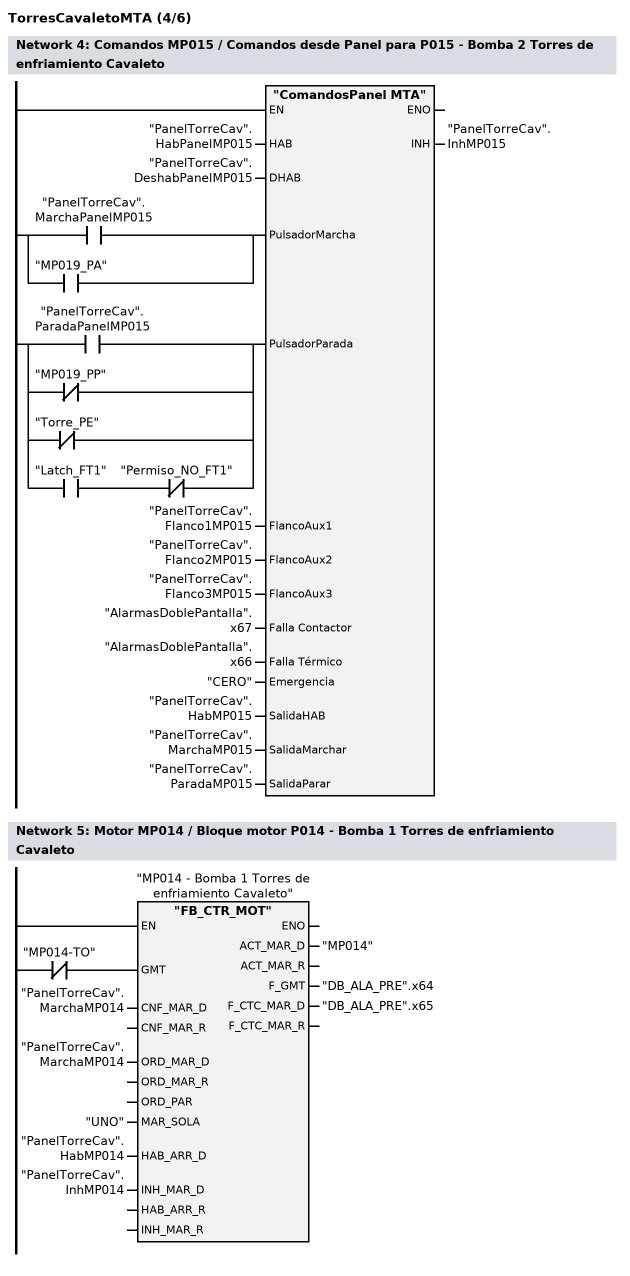
   RUNG wire#powerrail
      "ComandosPanel MTA"(PulsadorMarcha := wire#w1, PulsadorParada := wire#w2, HAB := "PanelTorreCav".HabPanelMP015, DHAB := "PanelTorreCav".DeshabPanelMP015, FlancoAux1 := "PanelTorreCav".Flanco1MP015, FlancoAux2 := "PanelTorreCav".Flanco2MP015, FlancoAux3 := "PanelTorreCav".Flanco3MP015, "Falla Contactor" := "AlarmasDoblePantalla".x67, "Falla Térmico" := "AlarmasDoblePantalla".x66, Emergencia := "CERO", SalidaHAB := "PanelTorreCav".HabMP015, SalidaMarchar := "PanelTorreCav".MarchaMP015, SalidaParar := "PanelTorreCav".ParadaMP015, INH => "PanelTorreCav".InhMP015)
   END_RUNG
   RUNG wire#powerrail
      Contact( "PanelTorreCav".MarchaPanelMP015 )
   END_RUNG wire#w1
   RUNG wire#powerrail
      Contact( "MP019_PA" )
   END_RUNG wire#w1
   RUNG wire#powerrail
      Contact( "PanelTorreCav".ParadaPanelMP015 )
   END_RUNG wire#w2
   RUNG wire#powerrail
      I_Contact( "MP019_PP" )
   END_RUNG wire#w2
   RUNG wire#powerrail
      I_Contact( "Torre_PE" )
   END_RUNG wire#w2
   RUNG wire#powerrail
      Contact( "Latch_FT1" )
      I_Contact( "Permiso_NO_FT1" )
   END_RUNG wire#w2
   // the same network as SCL:
   "ComandosPanel MTA"(HAB := "PanelTorreCav".HabPanelMP015,
                       DHAB := "PanelTorreCav".DeshabPanelMP015,
                       PulsadorMarcha := "PanelTorreCav".MarchaPanelMP015 OR "MP019_PA",
                       PulsadorParada := "PanelTorreCav".ParadaPanelMP015 OR NOT "MP019_PP" OR NOT "Torre_PE" OR ("Latch_FT1" AND NOT "Permiso_NO_FT1"),
                       FlancoAux1 := "PanelTorreCav".Flanco1MP015,
                       FlancoAux2 := "PanelTorreCav".Flanco2MP015,
                       FlancoAux3 := "PanelTorreCav".Flanco3MP015,
                       "Falla Contactor" := "AlarmasDoblePantalla".x67,
                       "Falla Térmico" := "AlarmasDoblePantalla".x66,
                       Emergencia := "CERO",
                       SalidaHAB := "PanelTorreCav".HabMP015,
                       SalidaMarchar := "PanelTorreCav".MarchaMP015,
                       SalidaParar := "PanelTorreCav".ParadaMP015,
                       INH => "PanelTorreCav".InhMP015);
END_REGION

REGION Network 5: Motor MP014 / Bloque motor P014 - Bomba 1 Torres de enfriamiento Cavaleto
   RUNG wire#powerrail
      "MP014 - Bomba 1 Torres de enfriamiento Cavaleto"(CNF_MAR_D := "PanelTorreCav".MarchaMP014, CNF_MAR_R :=, ORD_MAR_D := "PanelTorreCav".MarchaMP014, ORD_MAR_R :=, ORD_PAR :=, MAR_SOLA := "UNO", HAB_ARR_D := "PanelTorreCav".HabMP014, INH_MAR_D := "PanelTorreCav".InhMP014, HAB_ARR_R :=, INH_MAR_R :=, ACT_MAR_D => "MP014", ACT_MAR_R =>, F_GMT => "DB_ALA_PRE".x64, F_CTC_MAR_D => "DB_ALA_PRE".x65, F_CTC_MAR_R =>, GMT := wire#w1)
   END_RUNG
   RUNG wire#powerrail
      I_Contact( "MP014-TO" )
   END_RUNG wire#w1
   // the same network as SCL:
   "MP014 - Bomba 1 Torres de enfriamiento Cavaleto"(GMT := NOT "MP014-TO",   // "FB_CTR_MOT"
                           CNF_MAR_D := "PanelTorreCav".MarchaMP014,
                           ORD_MAR_D := "PanelTorreCav".MarchaMP014,
                           MAR_SOLA := "UNO",
                           HAB_ARR_D := "PanelTorreCav".HabMP014,
                           INH_MAR_D := "PanelTorreCav".InhMP014,
                           ACT_MAR_D => "MP014",
                           F_GMT => "DB_ALA_PRE".x64,
                           F_CTC_MAR_D => "DB_ALA_PRE".x65);
END_REGION

REGION Network 6: Motor MP015 / Bloque motor P015 - Bomba 2 Torres de enfriamiento Cavaleto
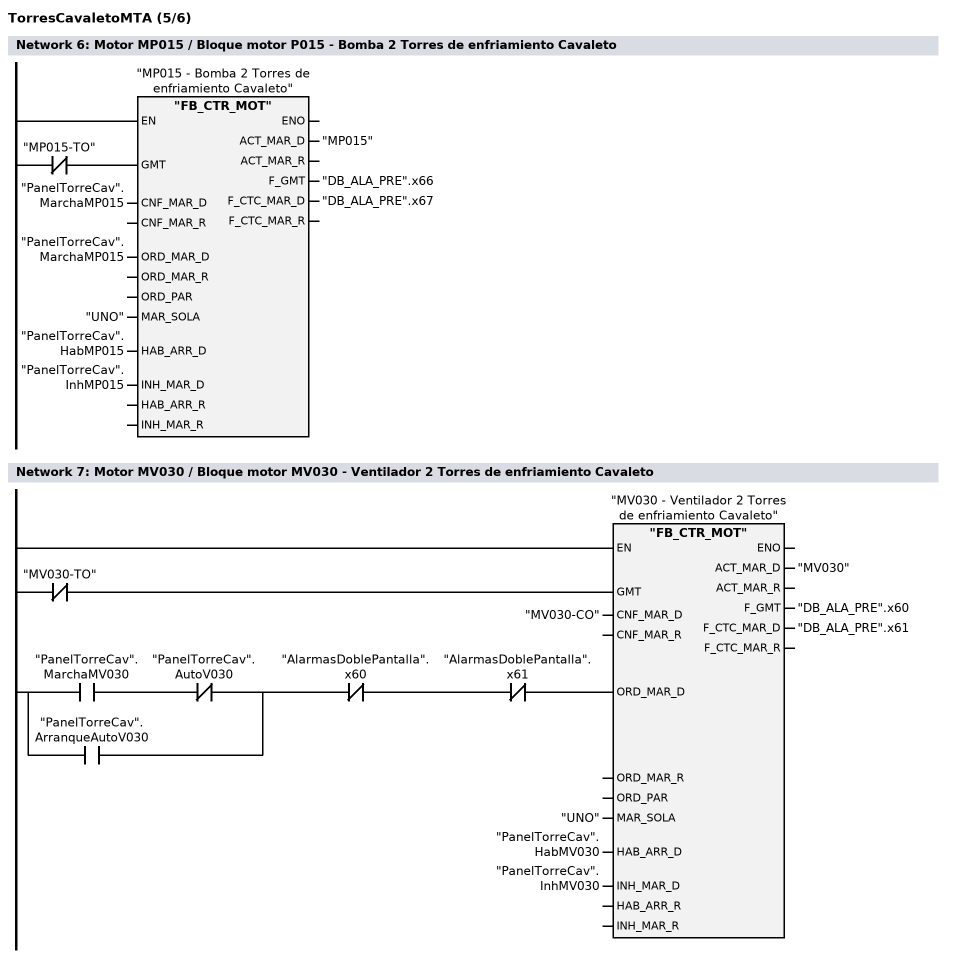
   RUNG wire#powerrail
      "MP015 - Bomba 2 Torres de enfriamiento Cavaleto"(CNF_MAR_D := "PanelTorreCav".MarchaMP015, CNF_MAR_R :=, ORD_MAR_D := "PanelTorreCav".MarchaMP015, ORD_MAR_R :=, ORD_PAR :=, MAR_SOLA := "UNO", HAB_ARR_D := "PanelTorreCav".HabMP015, INH_MAR_D := "PanelTorreCav".InhMP015, HAB_ARR_R :=, INH_MAR_R :=, ACT_MAR_D => "MP015", ACT_MAR_R =>, F_GMT => "DB_ALA_PRE".x66, F_CTC_MAR_D => "DB_ALA_PRE".x67, F_CTC_MAR_R =>, GMT := wire#w1)
   END_RUNG
   RUNG wire#powerrail
      I_Contact( "MP015-TO" )
   END_RUNG wire#w1
   // the same network as SCL:
   "MP015 - Bomba 2 Torres de enfriamiento Cavaleto"(GMT := NOT "MP015-TO",   // "FB_CTR_MOT"
                           CNF_MAR_D := "PanelTorreCav".MarchaMP015,
                           ORD_MAR_D := "PanelTorreCav".MarchaMP015,
                           MAR_SOLA := "UNO",
                           HAB_ARR_D := "PanelTorreCav".HabMP015,
                           INH_MAR_D := "PanelTorreCav".InhMP015,
                           ACT_MAR_D => "MP015",
                           F_GMT => "DB_ALA_PRE".x66,
                           F_CTC_MAR_D => "DB_ALA_PRE".x67);
END_REGION

REGION Network 7: Motor MV030 / Bloque motor MV030 - Ventilador 2 Torres de enfriamiento Cavaleto
   RUNG wire#powerrail
      "MV030 - Ventilador 2 Torres de enfriamiento Cavaleto"(GMT := wire#w1, ORD_MAR_D := wire#w3, CNF_MAR_D := "MV030-CO", CNF_MAR_R :=, ORD_MAR_R :=, ORD_PAR :=, MAR_SOLA := "UNO", HAB_ARR_D := "PanelTorreCav".HabMV030, INH_MAR_D := "PanelTorreCav".InhMV030, HAB_ARR_R :=, INH_MAR_R :=, ACT_MAR_D => "MV030", ACT_MAR_R =>, F_GMT => "DB_ALA_PRE".x60, F_CTC_MAR_D => "DB_ALA_PRE".x61, F_CTC_MAR_R =>)
   END_RUNG
   RUNG wire#powerrail
      I_Contact( "MV030-TO" )
   END_RUNG wire#w1
   RUNG wire#powerrail
      Contact( "PanelTorreCav".MarchaMV030 )
      I_Contact( "PanelTorreCav".AutoV030 )
      wire#w2
      I_Contact( "AlarmasDoblePantalla".x60 )
      I_Contact( "AlarmasDoblePantalla".x61 )
   END_RUNG wire#w3
   RUNG wire#powerrail
      Contact( "PanelTorreCav".ArranqueAutoV030 )
   END_RUNG wire#w2
   // the same network as SCL:
   "MV030 - Ventilador 2 Torres de enfriamiento Cavaleto"(GMT := NOT "MV030-TO",   // "FB_CTR_MOT"
                           CNF_MAR_D := "MV030-CO",
                           ORD_MAR_D := (("PanelTorreCav".MarchaMV030 AND NOT "PanelTorreCav".AutoV030) OR "PanelTorreCav".ArranqueAutoV030) AND NOT "AlarmasDoblePantalla".x60 AND NOT "AlarmasDoblePantalla".x61,
                           MAR_SOLA := "UNO",
                           HAB_ARR_D := "PanelTorreCav".HabMV030,
                           INH_MAR_D := "PanelTorreCav".InhMV030,
                           ACT_MAR_D => "MV030",
                           F_GMT => "DB_ALA_PRE".x60,
                           F_CTC_MAR_D => "DB_ALA_PRE".x61);
END_REGION

REGION Network 8: Motor MV031 / Bloque motorMV031 - Ventilador 1 Torres de enfriamiento Cavaleto
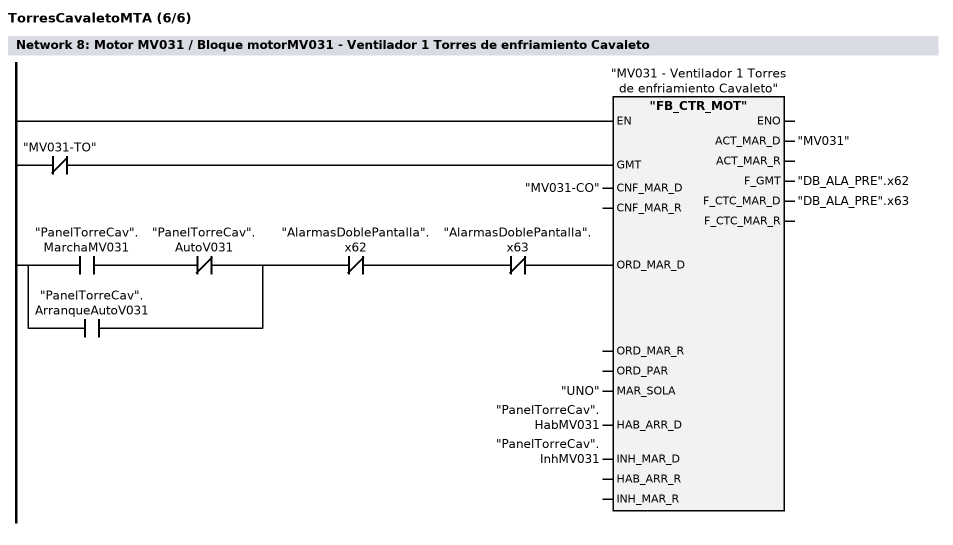
   RUNG wire#powerrail
      "MV031 - Ventilador 1 Torres de enfriamiento Cavaleto"(GMT := wire#w1, ORD_MAR_D := wire#w3, CNF_MAR_D := "MV031-CO", CNF_MAR_R :=, ORD_MAR_R :=, ORD_PAR :=, MAR_SOLA := "UNO", HAB_ARR_D := "PanelTorreCav".HabMV031, INH_MAR_D := "PanelTorreCav".InhMV031, HAB_ARR_R :=, INH_MAR_R :=, ACT_MAR_D => "MV031", ACT_MAR_R =>, F_GMT => "DB_ALA_PRE".x62, F_CTC_MAR_D => "DB_ALA_PRE".x63, F_CTC_MAR_R =>)
   END_RUNG
   RUNG wire#powerrail
      I_Contact( "MV031-TO" )
   END_RUNG wire#w1
   RUNG wire#powerrail
      Contact( "PanelTorreCav".MarchaMV031 )
      I_Contact( "PanelTorreCav".AutoV031 )
      wire#w2
      I_Contact( "AlarmasDoblePantalla".x62 )
      I_Contact( "AlarmasDoblePantalla".x63 )
   END_RUNG wire#w3
   RUNG wire#powerrail
      Contact( "PanelTorreCav".ArranqueAutoV031 )
   END_RUNG wire#w2
   // the same network as SCL:
   "MV031 - Ventilador 1 Torres de enfriamiento Cavaleto"(GMT := NOT "MV031-TO",   // "FB_CTR_MOT"
                           CNF_MAR_D := "MV031-CO",
                           ORD_MAR_D := (("PanelTorreCav".MarchaMV031 AND NOT "PanelTorreCav".AutoV031) OR "PanelTorreCav".ArranqueAutoV031) AND NOT "AlarmasDoblePantalla".x62 AND NOT "AlarmasDoblePantalla".x63,
                           MAR_SOLA := "UNO",
                           HAB_ARR_D := "PanelTorreCav".HabMV031,
                           INH_MAR_D := "PanelTorreCav".InhMV031,
                           ACT_MAR_D => "MV031",
                           F_GMT => "DB_ALA_PRE".x62,
                           F_CTC_MAR_D => "DB_ALA_PRE".x63);
END_REGION
END_FUNCTION

// folder: Torres de Agua/Torres Chillers

FUNCTION "TorresAutoMTA" : Void   // FC9, LAD
{ S7_Optimized_Access := 'FALSE' }
VERSION : 0.1
   VAR_TEMP
      TEMP0 : DInt;
   END_VAR
BEGIN

REGION Network 1: Lectura Temperatura de Torres Chillers
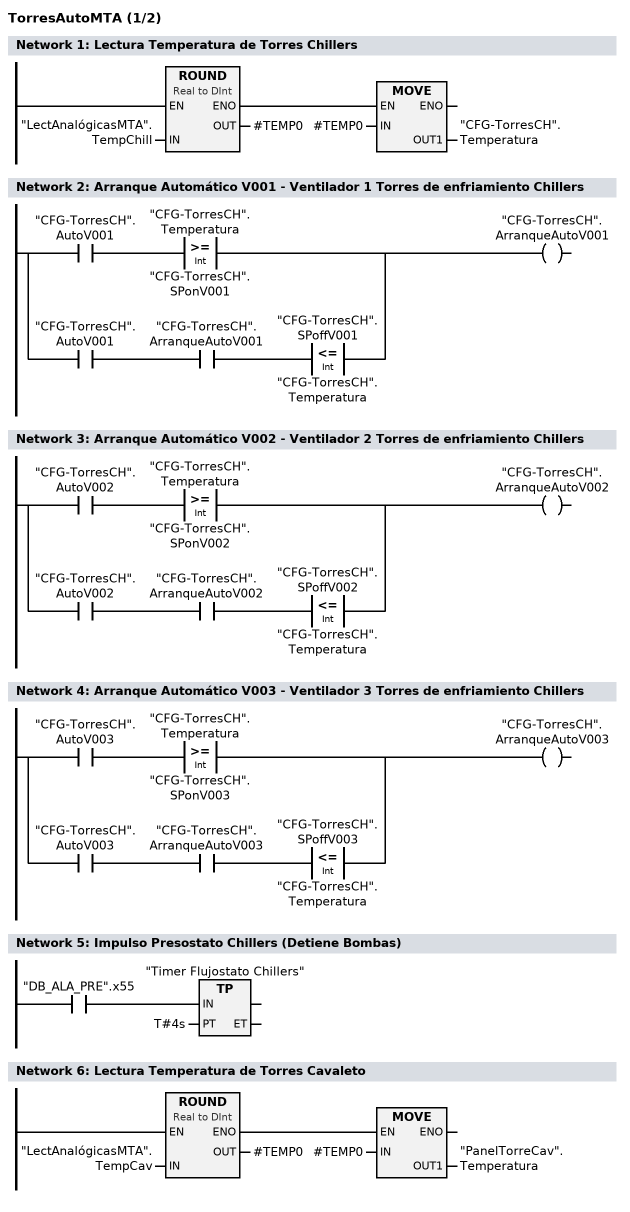
   RUNG wire#powerrail
      { S7_Templates := "[SrcType := Real, DestType := DInt]"; S7_GenerateENO := "TRUE" } Round(in := "LectAnalógicasMTA".TempChill, out => #TEMP0)
      { S7_GenerateENO := "TRUE" } Move(in := #TEMP0, out1 => "CFG-TorresCH".Temperatura)
   END_RUNG
   // the same network as SCL:
   // ENO of a box is taken as its EN; it also drops when the box reports an error
   #TEMP0 := ROUND("LectAnalógicasMTA".TempChill);
   "CFG-TorresCH".Temperatura := #TEMP0;
END_REGION

REGION Network 2: Arranque Automático V001 - Ventilador 1 Torres de enfriamiento Chillers
   RUNG wire#powerrail
      Contact( "CFG-TorresCH".AutoV001 )
      { S7_Templates := "SrcType := Int" } GE_Contact(in1 := "CFG-TorresCH".Temperatura, in2 := "CFG-TorresCH".SPonV001)
      wire#w1
      Coil( "CFG-TorresCH".ArranqueAutoV001 )
   END_RUNG
   RUNG wire#powerrail
      Contact( "CFG-TorresCH".AutoV001 )
      Contact( "CFG-TorresCH".ArranqueAutoV001 )
      { S7_Templates := "SrcType := Int" } LE_Contact(in1 := "CFG-TorresCH".SPoffV001, in2 := "CFG-TorresCH".Temperatura)
   END_RUNG wire#w1
   // the same network as SCL:
   "CFG-TorresCH".ArranqueAutoV001 := ("CFG-TorresCH".AutoV001 AND ("CFG-TorresCH".Temperatura >= "CFG-TorresCH".SPonV001)) OR ("CFG-TorresCH".AutoV001 AND "CFG-TorresCH".ArranqueAutoV001 AND ("CFG-TorresCH".SPoffV001 <= "CFG-TorresCH".Temperatura));
END_REGION

REGION Network 3: Arranque Automático V002 - Ventilador 2 Torres de enfriamiento Chillers
   RUNG wire#powerrail
      Contact( "CFG-TorresCH".AutoV002 )
      { S7_Templates := "SrcType := Int" } GE_Contact(in1 := "CFG-TorresCH".Temperatura, in2 := "CFG-TorresCH".SPonV002)
      wire#w1
      Coil( "CFG-TorresCH".ArranqueAutoV002 )
   END_RUNG
   RUNG wire#powerrail
      Contact( "CFG-TorresCH".AutoV002 )
      Contact( "CFG-TorresCH".ArranqueAutoV002 )
      { S7_Templates := "SrcType := Int" } LE_Contact(in1 := "CFG-TorresCH".SPoffV002, in2 := "CFG-TorresCH".Temperatura)
   END_RUNG wire#w1
   // the same network as SCL:
   "CFG-TorresCH".ArranqueAutoV002 := ("CFG-TorresCH".AutoV002 AND ("CFG-TorresCH".Temperatura >= "CFG-TorresCH".SPonV002)) OR ("CFG-TorresCH".AutoV002 AND "CFG-TorresCH".ArranqueAutoV002 AND ("CFG-TorresCH".SPoffV002 <= "CFG-TorresCH".Temperatura));
END_REGION

REGION Network 4: Arranque Automático V003 - Ventilador 3 Torres de enfriamiento Chillers
   RUNG wire#powerrail
      Contact( "CFG-TorresCH".AutoV003 )
      { S7_Templates := "SrcType := Int" } GE_Contact(in1 := "CFG-TorresCH".Temperatura, in2 := "CFG-TorresCH".SPonV003)
      wire#w1
      Coil( "CFG-TorresCH".ArranqueAutoV003 )
   END_RUNG
   RUNG wire#powerrail
      Contact( "CFG-TorresCH".AutoV003 )
      Contact( "CFG-TorresCH".ArranqueAutoV003 )
      { S7_Templates := "SrcType := Int" } LE_Contact(in1 := "CFG-TorresCH".SPoffV003, in2 := "CFG-TorresCH".Temperatura)
   END_RUNG wire#w1
   // the same network as SCL:
   "CFG-TorresCH".ArranqueAutoV003 := ("CFG-TorresCH".AutoV003 AND ("CFG-TorresCH".Temperatura >= "CFG-TorresCH".SPonV003)) OR ("CFG-TorresCH".AutoV003 AND "CFG-TorresCH".ArranqueAutoV003 AND ("CFG-TorresCH".SPoffV003 <= "CFG-TorresCH".Temperatura));
END_REGION

REGION Network 5: Impulso Presostato Chillers (Detiene Bombas)
   "Timer Flujostato Chillers".TP(IN := "DB_ALA_PRE".x55, PT := T#4s);
END_REGION

REGION Network 6: Lectura Temperatura de Torres Cavaleto
   RUNG wire#powerrail
      { S7_Templates := "[SrcType := Real, DestType := DInt]"; S7_GenerateENO := "TRUE" } Round(in := "LectAnalógicasMTA".TempCav, out => #TEMP0)
      { S7_GenerateENO := "TRUE" } Move(in := #TEMP0, out1 => "PanelTorreCav".Temperatura)
   END_RUNG
   // the same network as SCL:
   // ENO of a box is taken as its EN; it also drops when the box reports an error
   #TEMP0 := ROUND("LectAnalógicasMTA".TempCav);
   "PanelTorreCav".Temperatura := #TEMP0;
END_REGION

REGION Network 7: Arranque Automático MV030 - Ventilador 1 Torres de enfriamiento Cavaleto
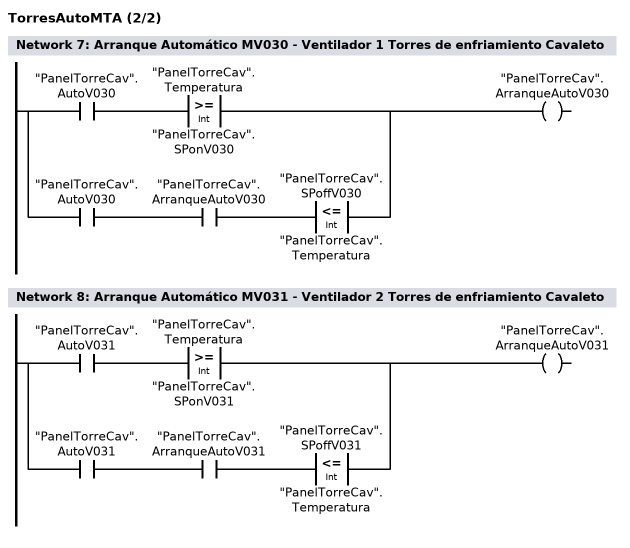
   RUNG wire#powerrail
      Contact( "PanelTorreCav".AutoV030 )
      { S7_Templates := "SrcType := Int" } GE_Contact(in1 := "PanelTorreCav".Temperatura, in2 := "PanelTorreCav".SPonV030)
      wire#w1
      Coil( "PanelTorreCav".ArranqueAutoV030 )
   END_RUNG
   RUNG wire#powerrail
      Contact( "PanelTorreCav".AutoV030 )
      Contact( "PanelTorreCav".ArranqueAutoV030 )
      { S7_Templates := "SrcType := Int" } LE_Contact(in1 := "PanelTorreCav".SPoffV030, in2 := "PanelTorreCav".Temperatura)
   END_RUNG wire#w1
   // the same network as SCL:
   "PanelTorreCav".ArranqueAutoV030 := ("PanelTorreCav".AutoV030 AND ("PanelTorreCav".Temperatura >= "PanelTorreCav".SPonV030)) OR ("PanelTorreCav".AutoV030 AND "PanelTorreCav".ArranqueAutoV030 AND ("PanelTorreCav".SPoffV030 <= "PanelTorreCav".Temperatura));
END_REGION

REGION Network 8: Arranque Automático MV031 - Ventilador 2 Torres de enfriamiento Cavaleto
   RUNG wire#powerrail
      Contact( "PanelTorreCav".AutoV031 )
      { S7_Templates := "SrcType := Int" } GE_Contact(in1 := "PanelTorreCav".Temperatura, in2 := "PanelTorreCav".SPonV031)
      wire#w1
      Coil( "PanelTorreCav".ArranqueAutoV031 )
   END_RUNG
   RUNG wire#powerrail
      Contact( "PanelTorreCav".AutoV031 )
      Contact( "PanelTorreCav".ArranqueAutoV031 )
      { S7_Templates := "SrcType := Int" } LE_Contact(in1 := "PanelTorreCav".SPoffV031, in2 := "PanelTorreCav".Temperatura)
   END_RUNG wire#w1
   // the same network as SCL:
   "PanelTorreCav".ArranqueAutoV031 := ("PanelTorreCav".AutoV031 AND ("PanelTorreCav".Temperatura >= "PanelTorreCav".SPonV031)) OR ("PanelTorreCav".AutoV031 AND "PanelTorreCav".ArranqueAutoV031 AND ("PanelTorreCav".SPoffV031 <= "PanelTorreCav".Temperatura));
END_REGION
END_FUNCTION

(* ===== HMI "HMI_RT_3" =====
system functions are stored by id; their names below are inferred from use
connection "Conexión2-PLC_1": ETHERNET, SIMATIC S7 300/400 MPI

HMI tags "AlarmasMTA"
   "AlarmasWord0" : Int AT %DB86.DBW0, 1 s
   "AlarmasWord1" : Int AT %DB86.DBW2, 1 s
   "AlarmasWord2" : Int AT %DB86.DBW4, 1 s
   "AlarmasWord3" : Int AT %DB86.DBW6, 1 s
   "AlarmasWord4" : Int AT %DB86.DBW8, 1 s
   "AlarmasWord5" : Int AT %DB86.DBW10, 1 s
   "AlarmasWord6" : Int AT %DB86.DBW12, 1 s
   "AlarmasWord7" : Int AT %DB86.DBW14, 1 s
   "AlarmasWord8" : Int AT %DB86.DBW16, 1 s
   "Rec0" : Int AT %DB86.DBW0, 1 s
   "Rec1" : Int AT %DB86.DBW2, 1 s
   "Rec2" : Int AT %DB86.DBW4, 1 s
   "Rec3" : Int AT %DB86.DBW6, 1 s
   "Rec4" : Int AT %DB86.DBW8, 1 s
   "Rec5" : Int AT %DB86.DBW10, 1 s
   "Rec6" : Int AT %DB86.DBW12, 1 s
   "Rec7" : Int AT %DB86.DBW14, 1 s
   "Rec8" : Int AT %DB86.DBW16, 1 s
   "AlarmasWord9" : Int AT %DB86.DBW18, 1 s
   "AlarmasWord10" : Int AT %DB86.DBW20, 1 s
   "AlarmasWord11" : Int AT %DB86.DBW22, 1 s
   "AlarmasWord12" : Int AT %DB86.DBW24, 1 s
   "AlarmasWord13" : Int AT %DB86.DBW26, 1 s
   "AlarmasWord14" : Int AT %DB86.DBW28, 1 s
   "Rec9" : Int AT %DB86.DBW18, 1 s
   "Rec10" : Int AT %DB86.DBW20, 1 s
   "Rec11" : Int AT %DB86.DBW22, 1 s
   "Rec12" : Int AT %DB86.DBW24, 1 s
   "Rec13" : Int AT %DB86.DBW26, 1 s
   "Rec14" : Int AT %DB86.DBW28, 1 s
   "AlarmasWord1(1)" : Int AT %DB86.DBW2, 1 s
   "AlarmasWord15" : Int AT %DB86.DBW30, 1 s
   "Rec15" : Int AT %DB86.DBW30, 1 s
   "EncendidoPLC" : Bool AT %M300.1, 1 s

HMI tags "AutoTorresChillers"
   "AutoV001" : Bool AT %DB92.DBX0.0, 1 s
   "AutoV002" : Bool AT %DB92.DBX0.1, 1 s
   "AutoV003" : Bool AT %DB92.DBX0.2, 1 s
   "SP-ON-V001" : Int AT %DB92.DBW2, 1 s
   "SP-ON-V002" : Int AT %DB92.DBW4, 1 s
   "SP-ON-V003" : Int AT %DB92.DBW6, 1 s
   "SP-OFF-V001" : Int AT %DB92.DBW8, 1 s
   "SP-OFF-V002" : Int AT %DB92.DBW10, 1 s
   "SP-OFF-V003" : Int AT %DB92.DBW12, 1 s
   "TemperaturatorresCH" : Real AT %DB52.DBD4, 1 s

HMI tags "CFG-Analog-MTA"
   "PresiónALTA" : Real AT %DB52.DBD52, 1 s
   "PresiónBAJA" : Real AT %DB52.DBD16, 1 s
   "TempCAV" : Real AT %DB52.DBD0, 1 s
   "TempCH" : Real AT %DB52.DBD4, 1 s
   "CFG-ALtaHH" : Real AT %DB52.DBD20, 1 s
   "CFG-ALtaH" : Real AT %DB52.DBD24, 1 s
   "CFG-ALtaL" : Real AT %DB52.DBD28, 1 s
   "CFG-ALtaLL" : Real AT %DB52.DBD32, 1 s
   "CFG-BajaHH" : Real AT %DB52.DBD36, 1 s
   "CFG-BajaH" : Real AT %DB52.DBD40, 1 s
   "CFG-BajaL" : Real AT %DB52.DBD44, 1 s
   "CFG-BajaLL" : Real AT %DB52.DBD48, 1 s

HMI tags "ChillersMTA"
   "HabMT007" : Bool AT %DB90.DBX6.4, 1 s
   "HabMT008" : Bool AT %DB90.DBX6.5, 1 s
   "HabMT009" : Bool AT %DB90.DBX6.6, 1 s
   "HabMT010" : Bool AT %DB90.DBX6.7, 1 s
   "DesMT007" : Bool AT %DB90.DBX8.1, 1 s
   "DesMT008" : Bool AT %DB90.DBX8.2, 1 s
   "DesMT009" : Bool AT %DB90.DBX8.3, 1 s
   "DesMT010" : Bool AT %DB90.DBX8.4, 1 s
   "MarchaMT007" : Bool AT %DB90.DBX9.6, 1 s
   "MarchaMT008" : Bool AT %DB90.DBX9.7, 1 s
   "MarchaMT009" : Bool AT %DB90.DBX10.0, 1 s
   "MarchaMT010" : Bool AT %DB90.DBX10.1, 1 s
   "ParadaMT007" : Bool AT %DB90.DBX11.3, 1 s
   "ParadaMT008" : Bool AT %DB90.DBX11.4, 1 s
   "ParadaMT009" : Bool AT %DB90.DBX11.5, 1 s
   "ParadaMT010" : Bool AT %DB90.DBX11.6, 1 s
   "Habilitación-CH-SOP-GR" : Bool AT %Q69.4, 1 s
   "Habilitación-CH-SOP-CH" : Bool AT %Q69.5, 1 s
   "Habilitación-CH-ENV-GR" : Bool AT %Q69.6, 1 s
   "Habilitación-CH-ENV-CH" : Bool AT %Q69.7, 1 s
   "Alarma1-CH-SOP-GR" : Bool AT %I68.4, 1 s
   "Alarma2-CH-SOP-GR" : Bool AT %I68.5, 1 s
   "RUN-CH-SOP-GR" : Bool AT %I68.6, 1 s
   "MAX-CH-SOP-GR" : Bool AT %I68.7, 1 s
   "AnimaciónMT007" : Byte AT %DB46.DBB6, 1 s
   "AnimaciónMT008" : Byte AT %DB46.DBB7, 1 s
   "AnimaciónMT009" : Byte AT %DB46.DBB8, 1 s
   "AnimaciónMT010" : Byte AT %DB46.DBB9, 1 s
   "AnimaciónMP010" : Byte AT %DB46.DBB0, 1 s
   "AnimaciónMP011" : Byte AT %DB46.DBB1, 1 s
   "AnimaciónMP012" : Byte AT %DB46.DBB2, 1 s
   "AnimaciónMP013" : Byte AT %DB46.DBB3, 1 s
   "HabMP010" : Bool AT %DB90.DBX7.0, 1 s
   "HabMP011" : Bool AT %DB90.DBX7.1, 1 s
   "HabMP012" : Bool AT %DB90.DBX7.2, 1 s
   "HabMP013" : Bool AT %DB90.DBX7.3, 1 s
   "HabMP018" : Bool AT %DB90.DBX7.4, 1 s
   "HabMP019" : Bool AT %DB90.DBX7.5, 1 s
   "DesMP010" : Bool AT %DB90.DBX8.5, 1 s
   "DesMP011" : Bool AT %DB90.DBX8.6, 1 s
   "DesMP012" : Bool AT %DB90.DBX8.7, 1 s
   "DesMP013" : Bool AT %DB90.DBX9.0, 1 s
   "DesMP018" : Bool AT %DB90.DBX9.1, 1 s
   "DesMP019" : Bool AT %DB90.DBX9.2, 1 s
   "MarchaMP010" : Bool AT %DB90.DBX10.2, 1 s
   "MarchaMP011" : Bool AT %DB90.DBX10.3, 1 s
   "MarchaMP012" : Bool AT %DB90.DBX10.4, 1 s
   "MarchaMP013" : Bool AT %DB90.DBX10.5, 1 s
   "MarchaMP018" : Bool AT %DB90.DBX10.6, 1 s
   "MarchaMP019" : Bool AT %DB90.DBX10.7, 1 s
   "ParadaMP010" : Bool AT %DB90.DBX11.7, 1 s
   "ParadaMP011" : Bool AT %DB90.DBX12.0, 1 s
   "ParadaMP012" : Bool AT %DB90.DBX12.1, 1 s
   "ParadaMP013" : Bool AT %DB90.DBX12.2, 1 s
   "ParadaMP018" : Bool AT %DB90.DBX12.3, 1 s
   "ParadaMP019" : Bool AT %DB90.DBX12.4, 1 s
   "AnimaciónMP018" : Byte AT %DB46.DBB4, 1 s
   "AnimaciónMP019" : Byte AT %DB46.DBB5, 1 s
   "DesV001" : Bool AT %DB90.DBX9.3, 1 s
   "DesV002" : Bool AT %DB90.DBX9.4, 1 s
   "HabV001" : Bool AT %DB90.DBX7.6, 1 s
   "HabV002" : Bool AT %DB90.DBX7.7, 1 s
   "MarchaV001" : Bool AT %DB90.DBX11.0, 1 s
   "MarchaV002" : Bool AT %DB90.DBX11.1, 1 s
   "ParadaV001" : Bool AT %DB90.DBX12.5, 1 s
   "ParadaV002" : Bool AT %DB90.DBX12.6, 1 s
   "AnimaciónV001" : Byte AT %DB46.DBB10, 1 s
   "AnimaciónV002" : Byte AT %DB46.DBB11, 1 s
   "VentiladoresMTA" : Bool, internal
   "MAX-CH-ENV-GR" : Bool AT %I69.7, 1 s
   "RUN-CH-ENV-GR" : Bool AT %I69.6, 1 s
   "Alarma2-CH-ENV-GR" : Bool AT %I69.5, 1 s
   "Alarma1-CH-ENV-GR" : Bool AT %I69.4, 1 s
   "SirenaM1" : Bool AT %DB91.DBX0.0, 1 s
   "SirenaM2" : Bool AT %DB91.DBX0.1, 1 s
   "SirenaM3" : Bool AT %DB91.DBX0.2, 1 s
   "SirenaM4" : Bool AT %DB91.DBX0.3, 1 s
   "AnimaciónV003" : Byte AT %DB46.DBB12, 1 s
   "HabV003" : Bool AT %DB90.DBX8.0, 1 s
   "DesV003" : Bool AT %DB90.DBX9.5, 1 s
   "MarchaV003" : Bool AT %DB90.DBX11.2, 1 s
   "ParadaV003" : Bool AT %DB90.DBX12.7, 1 s
   "BombaTorreON" : Bool AT %M69.2, 1 s
   "SirenaM5" : Bool AT %DB91.DBX0.4, 1 s
   "SirenaChillers" : Bool AT %Q68.1, 1 s
   "SirenaM6" : Bool AT %DB91.DBX0.5, 1 s
   "SirenaM7" : Bool AT %DB91.DBX0.6, 1 s
   "SirenaM8" : Bool AT %DB91.DBX0.7, 1 s
   "SirenaM9" : Bool AT %DB91.DBX1.0, 1 s
   "SirenaM10" : Bool AT %DB91.DBX1.1, 1 s
   "AlarmaNueva" : Bool AT %DB47.DBX0.0, 1 s
   "AlarmaPresente" : Bool AT %DB47.DBX0.1, 1 s
   "SinAlarmas" : Bool AT %DB47.DBX0.2, 1 s
   "AlarmaAceite-CH-ENV-CH" : Bool AT %I76.0, 1 s
   "AlarmaTemp-CH-ENV-CH" : Bool AT %I76.1, 1 s
   "RUN-CH-ENV-CH" : Bool AT %I76.2, 1 s
   "VerCh1MTA" : Bool, internal
   "VerCh2MTA" : Bool, internal
   "VerCh3MTA" : Bool, internal
   "VerCh4MTA" : Bool, internal
   "AlarmaPRUEBA" : DWord AT %DB1.DBD0, 1 s
   "Presosato" : Bool AT %I76.4, 1 s
   "CH-SOP-CH-CTC1ON" : Bool AT %I69.0, 1 s
   "CH-SOP-CH-CTC2ON" : Bool AT %I69.1, 1 s
   "CH-SOP-CH-TERM1" : Bool AT %I69.2, 1 s
   "CH-SOP-CH-TERM2" : Bool AT %I69.3, 1 s
   "CH-ENV-CH-ACT" : Bool AT %I76.0, 1 s
   "CH-ENV-CH-TEMP" : Bool AT %I76.1, 1 s
   "CH-ENV-CH-TERM" : Bool AT %I76.2, 1 s
   "CH-ENV-CH-RUN" : Bool AT %I76.3, 1 s
   "BombaTorreON2" : Bool AT %M69.3, 1 s
   "HabV001(1)" : Bool AT %DB90.DBX7.6, 1 s
   "HabV002(1)" : Bool AT %DB90.DBX7.7, 1 s
   "HabV003(1)" : Bool AT %DB90.DBX8.0, 1 s
   "HabV4" : Bool AT %DB90.DBX8.1, 1 s
   "MarchaV001(1)" : Bool AT %DB90.DBX11.0, 1 s
   "MarchaV002(1)" : Bool AT %DB90.DBX11.1, 1 s
   "MarchaV003(1)" : Bool AT %DB90.DBX11.2, 1 s
   "ParadaV001(1)" : Bool AT %DB90.DBX12.5, 1 s
   "ParadaV002(1)" : Bool AT %DB90.DBX12.6, 1 s
   "ParadaV003(1)" : Bool AT %DB90.DBX12.7, 1 s
   "AnimaMenuV001" : Int AT %DB46.DBW24, 1 s
   "AnimaMenuV002" : Int AT %DB46.DBW26, 1 s
   "AnimaMenuV003" : Int AT %DB46.DBW28, 1 s
   "DeshV001" : Bool AT %DB90.DBX9.3, 1 s
   "DeshV002" : Bool AT %DB90.DBX9.4, 1 s
   "DeshV003" : Bool AT %DB90.DBX9.5, 1 s

discrete alarms
   125: 'Falla Contactor - V001 - Ventilador 1 Torres de enfriamiento Chillers', class MTA, trigger "Rec4" bit 8
   126: 'Falla Guardamotor - V001 - Ventilador 1 Torres de enfriamiento Chillers', class MTA, trigger "Rec3" bit 15
   127: 'Falla Guardamotor - V003 - Ventilador 3 Torres de enfriamiento Chillers', class MTA, trigger "Rec4" bit 11
   128: 'Falla Contactor - V002 - Ventilador 2 Torres de enfriamiento Chillers', class MTA, trigger "Rec4" bit 10
   129: 'Falla Guardamotor - V002 - Ventilador 2 Torres de enfriamiento Chillers', class MTA, trigger "Rec4" bit 9
   130: 'Falla Guardamotor - MP018 - Bomba 1 Torres de enfriamiento Chillers', class MTA, trigger "Rec3" bit 11
   131: 'Falla Contactor - MP013 - Bomba Backup Ch. Envasado', class MTA, trigger "Rec3" bit 10
   132: 'Falla Guardamotor - MP013 - Bomba Backup Ch. Envasado', class MTA, trigger "Rec3" bit 9
   133: 'Falla Contactor - MP019 - Bomba 2 Torres de enfriamiento Chillers', class MTA, trigger "Rec3" bit 14
   134: 'Falla Guardamotor - MP019 - Bomba 2 Torres de enfriamiento Chillers', class MTA, trigger "Rec3" bit 13
   135: 'Falla Contactor - MP018 - Bomba 1 Torres de enfriamiento Chillers', class MTA, trigger "Rec3" bit 12
   136: 'Falla Contactor - V003 - Ventilador 3 Torres de enfriamiento Chillers', class MTA, trigger "Rec4" bit 12
   137: 'Falla Guardamotor - MC061 - Compresor de Baja SULLAIR 1', class MTA, trigger "Rec4" bit 15
   138: 'Falla Contactor - MC060 - Compresor de Baja SULLAIR 2', class MTA, trigger "Rec4" bit 14
   139: 'Falla Guardamotor - MC060 - Compresor de Baja SULLAIR 2', class MTA, trigger "Rec4" bit 13
   140: 'Falla Contactor - MP012 - Bomba Principal Ch. Envasado', class MTA, trigger "Rec3" bit 8
   141: 'Alarma Presente en Chiller de envasado Grande', class MTA, trigger "Rec1" bit 8
   144: 'Falla Guardamotor - MT007 - Sopladora Línea 1', class MTA, trigger "Rec1" bit 11
   145: 'Chiller de envasado Grande en su máxima capacidad', class MTA, trigger "Rec1" bit 10
   146: 'Chiller de soplado Grande en su máxima capacidad', class MTA, trigger "Rec1" bit 9
   153: 'Falla Contactor - MT007 -Sopladora Línea 1', class MTA, trigger "Rec1" bit 12
   154: 'Falla Contactor - MP010 - Bomba Principal Ch. Soplado', class MTA, trigger "Rec2" bit 12
   155: 'Falla Guardamotor - MP010 - Bomba Principal Ch. Soplado', class MTA, trigger "Rec2" bit 11
   156: 'Falla Contactor - MT010 - Bomba Int L1 y Manomec', class MTA, trigger "Rec2" bit 10
   157: 'Falla Guardamotor - MP012 - Bomba Principal Ch. Envasado', class MTA, trigger "Rec2" bit 15
   158: 'Falla Contactor - MP011 - Bomba Backup Ch. Soplado', class MTA, trigger "Rec2" bit 14
   159: 'Falla Guardamotor - MP011 - Bomba Backup Ch. Soplado', class MTA, trigger "Rec2" bit 13
   160: 'Falla Guardamotor - MT009 - Bomba Int. L3 y L5', class MTA, trigger "Rec1" bit 15
   161: 'Falla Contactor - MT008 - Sopladora Línea 3 y Man.', class MTA, trigger "Rec1" bit 14
   162: 'Falla Guardamotor - MT008 - Sopladora Línea 3 y Man.', class MTA, trigger "Rec1" bit 13
   163: 'Falla Guardamotor - MT010 - Bomba Int L1 y Manomec', class MTA, trigger "Rec2" bit 9
   164: 'Falla Contactor - MT009 - Bomba Int. L3 y L5', class MTA, trigger "Rec2" bit 8
   165: 'Falla Contactor - MC061 - Compresor de Baja SULLAIR 1', class MTA, trigger "Rec5" bit 8
   166: 'Falla Guardamotor - MC062 - Compresor de Baja SULLAIR 0', class MTA, trigger "Rec5" bit 9
   167: 'Falla Contactor - MC062 - Compresor de Baja SULLAIR 0', class MTA, trigger "Rec5" bit 10
   168: 'Falla Guardamotor - MC063 - Compresor de Baja ATLAS 3', class MTA, trigger "Rec5" bit 11
   169: 'Falla Contactor - MC063 - Compresor de Baja ATLAS 3', class MTA, trigger "Rec5" bit 12
   170: 'Falla Guardamotor - MC064 - Compresor de Baja ATLAS 2', class MTA, trigger "Rec5" bit 13
   171: 'Falla Contactor - MC064 - Compresor de Baja ATLAS 2', class MTA, trigger "Rec5" bit 14
   172: 'Falla Guardamotor - MS050 - Secador de Alta ABC1', class MTA, trigger "Rec5" bit 15
   13: 'Falla Contactor - MS050 - Secador de Alta ABC1', class MTA, trigger "Rec6" bit 8
   14: 'Falla Guardamotor - MS051 - Secador de Alta ABC3', class MTA, trigger "Rec6" bit 9
   50: 'Falla Contactor - MS051 - Secador de Alta ABC3', class MTA, trigger "Rec6" bit 10
   53: 'Falla Guardamotor - MS052 - Secador de Alta ABC2', class MTA, trigger "Rec6" bit 11
   87: 'Falla Contactor - MS052 - Secador de Alta ABC2', class MTA, trigger "Rec6" bit 12
   88: 'Falla Guardamotor - MS053 - Secador de Alta FARGON', class MTA, trigger "Rec6" bit 13
   89: 'Falla Contactor - MS053 - Secador de Alta FARGON', class MTA, trigger "Rec6" bit 14
   90: 'Falla Presostato Chillers', class MTA, trigger "Rec6" bit 15
   69: 'Falla Contactor MS055 - Secador de Baja SULLAIR 2', class MTA, trigger "Rec7" bit 11
   68: 'Falla Guardamotor MS055 - Secador de Baja SULLAIR 2', class MTA, trigger "Rec7" bit 10
   67: 'Falla Contactor MS054 - Secador de Baja SULLAIR 1', class MTA, trigger "Rec7" bit 9
   66: 'Falla Guardamotor MS054 - Secador de Baja SULLAIR 1', class MTA, trigger "Rec7" bit 8
   70: 'Falla Guardamotor - MV030 - Ventilador 1 Torres de enfriamiento Cavaleto', class MTA, trigger "Rec7" bit 12
   71: 'Falla Contactor - MV030 - Ventilador 1 Torres de enfriamiento Cavaleto', class MTA, trigger "Rec7" bit 13
   72: 'Falla Guardamotor - MV031 - Ventilador 2 Torres de enfriamiento Cavaleto', class MTA, trigger "Rec7" bit 14
   73: 'Falla Contactor - MV031 - Ventilador 2 Torres de enfriamiento Cavaleto', class MTA, trigger "Rec7" bit 15
   74: 'Falla Guardamotor - MP014 - Bomba 1 Torres de enfriamiento Cavaleto', class MTA, trigger "Rec8" bit 8
   75: 'Falla Contactor - MP014 - Bomba 1 Torres de enfriamiento Cavaleto', class MTA, trigger "Rec8" bit 9
   76: 'Falla Guardamotor - MP015 - Bomba 2 Torres de enfriamiento Cavaleto', class MTA, trigger "Rec8" bit 10
   77: 'Falla Contactor - MP015 - Bomba 2 Torres de enfriamiento Cavaleto', class MTA, trigger "Rec8" bit 11
   78: 'Falla Guardamotor - MC001 - Compresor de Alta ABC2', class MTA, trigger "Rec8" bit 12
   79: 'Falla Contactor - MC001 - Compresor de Alta ABC2', class MTA, trigger "Rec8" bit 13
   80: 'Falla Guardamotor - MC002 - Compresor de Alta ABC3', class MTA, trigger "Rec8" bit 14
   81: 'Falla Contactor - MC002 - Compresor de Alta ABC3', class MTA, trigger "Rec8" bit 15
   82: 'Falla Guardamotor - MC003 - Compresor de Alta BELLIS', class MTA, trigger "Rec9" bit 8
   83: 'Falla Contactor - MC003 - Compresor de Alta BELLIS', class MTA, trigger "Rec9" bit 9
   91: 'Falla Guardamotor - MC004 - Compresor de Alta ABC4', class MTA, trigger "Rec9" bit 10
   92: 'Falla Contactor - MC004 - Compresor de Alta ABC4', class MTA, trigger "Rec9" bit 11
   93: 'Falla Guardamotor - MC005 - Compresor de Alta ABC5', class MTA, trigger "Rec9" bit 12
   94: 'Falla Contactor - MC005 - Compresor de Alta ABC5', class MTA, trigger "Rec9" bit 13
   96: 'Falla Compresor ABC2 Baja Presion de Aceite', class MTA, trigger "Rec9" bit 15
   97: 'Falla Compresor ABC2 Baja Presion de Agua', class MTA, trigger "Rec10" bit 8
   98: 'Falla Compresor ABC2 Alta Temperatura de Aire', class MTA, trigger "Rec10" bit 9
   99: 'Falla Compresor ABC2 Alta Temperatura de agua', class MTA, trigger "Rec10" bit 10
   100: 'Falla Compresor ABC3 Baja Presion de Aceite', class MTA, trigger "Rec10" bit 11
   101: 'Falla Compresor ABC3 Baja Presion de Agua', class MTA, trigger "Rec10" bit 12
   102: 'Falla Compresor ABC3 Alta Temperatura de Aire', class MTA, trigger "Rec10" bit 13
   121: 'Falla Compresor ABC3 Alta Temperatura de agua', class MTA, trigger "Rec10" bit 14
   104: 'Falla Compresor ABC4 Baja Presion de Aceite', class MTA, trigger "Rec10" bit 15
   105: 'Falla Compresor ABC4 Alta Temperatura de Aire', class MTA, trigger "Rec11" bit 8
   106: 'Falla Compresor ABC4 Alta Temperatura de Aire', class MTA, trigger "Rec11" bit 9
   107: 'Falla Compresor ABC4 Alta Temperatura de agua', class MTA, trigger "Rec11" bit 10
   108: 'Falla Compresor ABC5 Baja Presion de Aceite', class MTA, trigger "Rec11" bit 11
   109: 'Falla Compresor ABC5 Alta Temperatura de Aire', class MTA, trigger "Rec11" bit 12
   110: 'Falla Compresor ABC5 Alta Temperatura de Aire', class MTA, trigger "Rec11" bit 13
   111: 'Falla Compresor ABC5 Alta Temperatura de agua', class MTA, trigger "Rec11" bit 14
   112: 'Falla Compresor Bellis & MHW28 Baja Presion Aceite', class MTA, trigger "Rec11" bit 15
   113: 'Falla Compresor Bellis & MHW28 Baja Presion de Agua', class MTA, trigger "Rec12" bit 8
   114: 'Falla Compresor Bellis & MHW28 Alta temperatura de Aire', class MTA, trigger "Rec12" bit 9
   115: 'Falla Compresor Bellis & MHW28 Alta temperatura de Agua', class MTA, trigger "Rec12" bit 10
   116: 'Falla Compresor Bellis & MHW28 Falla de Flujostato', class MTA, trigger "Rec12" bit 11
   117: 'Compresor ABC2 Requiere Marcha', class MTA, trigger "Rec12" bit 12
   118: 'Compresor ABC3 Requiere Marcha', class MTA, trigger "Rec12" bit 13
   119: 'Compresor Bellis Requiere Marcha', class MTA, trigger "Rec12" bit 14
   120: 'Compresor ABC4 Requiere Marcha', class MTA, trigger "Rec12" bit 15
   122: 'Compresor ABC5 Requiere Marcha', class MTA, trigger "Rec13" bit 8
   1: 'Falla Conexión con sensor de Temperatura torres de Cavaleto', class MTA, trigger "Rec13" bit 9
   2: 'Falla Conexión con sensor de Temperatura torres de Chillers', class MTA, trigger "Rec13" bit 10
   3: 'Falla Conexión con sensor de Presión de ALTA', class MTA, trigger "Rec13" bit 11
   4: 'Falla Conexión con sensor de Presión de ALTA redundante', class MTA, trigger "Rec13" bit 12
   5: 'Falla Conexión con sensor de Presión de Baja', class MTA, trigger "Rec13" bit 13
   6: 'Falla Presión de Alta en Límite Mínimo', class MTA, trigger "Rec13" bit 14
   7: 'Falla Presión de Alta en demasiado Baja', class MTA, trigger "Rec13" bit 15
   8: 'Falla Presión de Alta en demasiado Alta', class MTA, trigger "Rec14" bit 8
   9: 'Falla Presión de Alta en Límite Máximo', class MTA, trigger "Rec14" bit 9
   10: 'Falla Presión de Baja en Límite Mínimo', class MTA, trigger "Rec14" bit 10
   11: 'Falla Presión de Baja en demasiado Baja', class MTA, trigger "Rec14" bit 11
   12: 'Falla Presión de Baja en demasiado Alta', class MTA, trigger "Rec14" bit 12
   15: 'Falla Presión de Baja en Límite Máximo', class MTA, trigger "Rec14" bit 13
   16: 'Falla en chiller de envasado chico', class MTA, trigger "Rec14" bit 14
   17: 'Falla en chiller de soplado chico', class MTA, trigger "Rec14" bit 15
   95: 'Falla Flujostato Torres Caveleto', class MTA, trigger "Rec9" bit 14
   149: 'Ninguna bomba de intercambiador de soplado en marcha', class MTA, trigger "Rec0" bit 8
   142: 'Alarma Presente en Chiller de soplado Grande', class MTA, trigger "Rec0" bit 15
   143: 'Ningún chiller de envasado habilitado', class MTA, trigger "Rec0" bit 14
   152: 'Ninguna bomba de chillers de envasado en marcha', class MTA, trigger "Rec0" bit 11
   147: 'Ninguna bomba de intercambiador de envasado en marcha', class MTA, trigger "Rec0" bit 10
   148: 'Ninguna bomba de chillers de soplado en marcha', class MTA, trigger "Rec0" bit 9
   150: 'Ningún Chiller de soplado habilitado', class MTA, trigger "Rec0" bit 13
   151: 'Ninguna bomba de torre de enfiamiento de chillers en marcha', class MTA, trigger "Rec0" bit 12
   21: 'El Compresor ABC4 alcanzó la máxima cantidad de horas', class MTA, trigger "Rec15" bit 11
   22: 'El Compresor ABC5 alcanzó la máxima cantidad de horas', class MTA, trigger "Rec15" bit 12
   19: 'El Compresor ABC3 alcanzó la máxima cantidad de horas', class MTA, trigger "Rec15" bit 9
   20: 'El Compresor Bellis alcanzó la máxima cantidad de horas', class MTA, trigger "Rec15" bit 10
   23: 'Falla algún contactor en Booster 1', class MTA, trigger "Rec15" bit 13
   24: 'Falla algún guardamotor en Booster 1', class MTA, trigger "Rec15" bit 14
   25: 'Presión Alta en Booster', class MTA, trigger "Rec15" bit 15
   18: 'El Compresor ABC2 alcanzó la máxima cantidad de horas', class MTA, trigger "Rec15" bit 8

text list "EstadoMotor": 0 'Detenido'; 1 'En Marcha'; 2 'Arrancando'; 3 'Deteniéndose'; 4 'Espera para Arrancar'; 5 'Sobrecarga de Corriente'; 6 'Deshabilitado'; 7 'En Falla'

graphic list "Motor2": 0 'Motor2Dorado'; 1 'Motor2Verde_1'; 2 'Motor2VerdeOscuro'; 3 'Motor2Azul'; 4 'Motor2Celeste'; 5 'Motor2Amarillo'; 6 'Motor2Gris_1'; 7 'Motor2Rojo'

graphic list "MotorTorre": 0 'torreFINAL4C2_1'; 1 'torreFINAL4C2v_2'; 2 'torreFINAL4C2v_2'; 3 'torreFINAL4C2b'; 4 'torreFINAL4C2b'; 5 'torreFINAL4C2a_2'; 6 'torreFINAL4C2_1'; 7 'torreFINAL4C2_1'

graphic list "Indicador": 0 'indDorado'; 1 'indVerde'; 2 'indVerde_1'; 3 'indAZUL'; 4 'indCeleste'; 5 'indAmarillo'; 6 'indGris'; 7 'indRojo'

graphic list "Secador2": 0 'BaseSullChicoDorado_2'; 1 'BaseSullChico_5'; 2 'BaseSullChico_5'; 3 'BaseSullChicoAzul_2'; 4 'BaseSullChicoAzul_2'; 5 'BaseSullChicoAmarillo_2'; 6 'BaseSullChicoGris_2'; 7 'BaseSullChicoRojo_2'

graphic list "Secador3": 0 'BaseSullChicoDorado_3'; 1 'BaseSullChico_6'; 2 'BaseSullChico_6'; 3 'BaseSullChicoAzul_3'; 4 'BaseSullChicoAzul_3'; 5 'BaseSullChicoAmarillo_3'; 6 'BaseSullChicoGris_3'; 7 'BaseSullChicoRojo_3'

graphic list "Secador1": 0 'BaseSullChicoDorado_1'; 1 'BaseSullChico_4'; 2 'BaseSullChico_4'; 3 'BaseSullChicoAzul_1'; 4 'BaseSullChicoAzul_1'; 5 'BaseSullChicoAmarillo_1'; 6 'BaseSullChicoGris_1'; 7 'BaseSullChicoRojo_1'

screen "MTA-Avisos" 800x480, template "Plantilla_2"
   AlarmView "Visor de avisos_1" at 5,53 size 790x367
   TextField "Campo de texto_5" at 327,10 size 54x27; Text 'Avisos'